DATA_BLOCK "MessagePrefix"   // DB31604
TITLE = CPG_MessagePrefix
{ S7_Optimized_Access := 'TRUE' }
AUTHOR : tech.team.motioncontrol@siemens.com
FAMILY : CPG
VERSION : 1.0
// Support: tech.team.motioncontrol@siemens.com
// Fax: +49 (0) 9131/98-1297
   VAR
      UN : Struct   // MessagePrefix for Unit
         Alarm : "CPG_typeMessagePrefix";   // MessagePrefix for Unit Alarms
      END_STRUCT;
      EM00 : Struct   // MessagePrefix for EquipmentModuleEM00
         EventControl : "CPG_typeMessagePrefix";   // MessagePrefixforEventControl
         CM01 : "CPG_typeMessagePrefix";   // MessagePrefixforControlModule#01
         CM02 : "CPG_typeMessagePrefix";   // MessagePrefixforControlModule#02
         CM03 : "CPG_typeMessagePrefix";   // MessagePrefixforControlModule#03
         CM04 : "CPG_typeMessagePrefix";   // MessagePrefixforControlModule#04
         CM05 : "CPG_typeMessagePrefix";   // MessagePrefixforControlModule#05
         CM06 : "CPG_typeMessagePrefix";   // MessagePrefixforControlModule#06
         CM07 : "CPG_typeMessagePrefix";   // MessagePrefixforControlModule#07
         CM08 : "CPG_typeMessagePrefix";   // MessagePrefixforControlModule#08
         CM09 : "CPG_typeMessagePrefix";   // MessagePrefixforControlModule#09
         CM10 : "CPG_typeMessagePrefix";   // MessagePrefixforControlModule#10
      END_STRUCT;
      EM01 : Struct   // MessagePrefix for EquipmentModuleEM01
         EventControl : "CPG_typeMessagePrefix";   // MessagePrefixforEventControl
         CM01 : "CPG_typeMessagePrefix";   // MessagePrefixforControlModule#01
         CM02 : "CPG_typeMessagePrefix";   // MessagePrefixforControlModule#02
         CM03 : "CPG_typeMessagePrefix";   // MessagePrefixforControlModule#03
         CM04 : "CPG_typeMessagePrefix";   // MessagePrefixforControlModule#04
         CM05 : "CPG_typeMessagePrefix";   // MessagePrefixforControlModule#05
         CM06 : "CPG_typeMessagePrefix";   // MessagePrefixforControlModule#06
         CM07 : "CPG_typeMessagePrefix";   // MessagePrefixforControlModule#07
         CM08 : "CPG_typeMessagePrefix";   // MessagePrefixforControlModule#08
         CM09 : "CPG_typeMessagePrefix";   // MessagePrefixforControlModule#09
         CM10 : "CPG_typeMessagePrefix";   // MessagePrefixforControlModule#10
      END_STRUCT;
      EM02 : Struct   // MessagePrefix for EquipmentModuleEM02
         EventControl : "CPG_typeMessagePrefix";   // MessagePrefixforEventControl
         CM01 : "CPG_typeMessagePrefix";   // MessagePrefixforControlModule#01
         CM02 : "CPG_typeMessagePrefix";   // MessagePrefixforControlModule#02
         CM03 : "CPG_typeMessagePrefix";   // MessagePrefixforControlModule#03
         CM04 : "CPG_typeMessagePrefix";   // MessagePrefixforControlModule#04
         CM05 : "CPG_typeMessagePrefix";   // MessagePrefixforControlModule#05
         CM06 : "CPG_typeMessagePrefix";   // MessagePrefixforControlModule#06
         CM07 : "CPG_typeMessagePrefix";   // MessagePrefixforControlModule#07
         CM08 : "CPG_typeMessagePrefix";   // MessagePrefixforControlModule#08
         CM09 : "CPG_typeMessagePrefix";   // MessagePrefixforControlModule#09
         CM10 : "CPG_typeMessagePrefix";   // MessagePrefixforControlModule#10
      END_STRUCT;
      EM03 : Struct   // MessagePrefix for EquipmentModuleEM03
         EventControl : "CPG_typeMessagePrefix";   // MessagePrefixforEventControl
         CM01 : "CPG_typeMessagePrefix";   // MessagePrefixforControlModule#01
         CM02 : "CPG_typeMessagePrefix";   // MessagePrefixforControlModule#02
         CM03 : "CPG_typeMessagePrefix";   // MessagePrefixforControlModule#03
         CM04 : "CPG_typeMessagePrefix";   // MessagePrefixforControlModule#04
         CM05 : "CPG_typeMessagePrefix";   // MessagePrefixforControlModule#05
         CM06 : "CPG_typeMessagePrefix";   // MessagePrefixforControlModule#06
         CM07 : "CPG_typeMessagePrefix";   // MessagePrefixforControlModule#07
         CM08 : "CPG_typeMessagePrefix";   // MessagePrefixforControlModule#08
         CM09 : "CPG_typeMessagePrefix";   // MessagePrefixforControlModule#09
         CM10 : "CPG_typeMessagePrefix";   // MessagePrefixforControlModule#10
      END_STRUCT;
      EM04 : Struct   // MessagePrefix for EquipmentModuleEM04
         EventControl : "CPG_typeMessagePrefix";   // MessagePrefixforEventControl
         CM01 : "CPG_typeMessagePrefix";   // MessagePrefixforControlModule#01
         CM02 : "CPG_typeMessagePrefix";   // MessagePrefixforControlModule#02
         CM03 : "CPG_typeMessagePrefix";   // MessagePrefixforControlModule#03
         CM04 : "CPG_typeMessagePrefix";   // MessagePrefixforControlModule#04
         CM05 : "CPG_typeMessagePrefix";   // MessagePrefixforControlModule#05
         CM06 : "CPG_typeMessagePrefix";   // MessagePrefixforControlModule#06
         CM07 : "CPG_typeMessagePrefix";   // MessagePrefixforControlModule#07
         CM08 : "CPG_typeMessagePrefix";   // MessagePrefixforControlModule#08
         CM09 : "CPG_typeMessagePrefix";   // MessagePrefixforControlModule#09
         CM10 : "CPG_typeMessagePrefix";   // MessagePrefixforControlModule#10
      END_STRUCT;
      EM05 : Struct   // MessagePrefix for EquipmentModuleEM05
         EventControl : "CPG_typeMessagePrefix";   // MessagePrefixforEventControl
         CM01 : "CPG_typeMessagePrefix";   // MessagePrefixforControlModule#01
         CM02 : "CPG_typeMessagePrefix";   // MessagePrefixforControlModule#02
         CM03 : "CPG_typeMessagePrefix";   // MessagePrefixforControlModule#03
         CM04 : "CPG_typeMessagePrefix";   // MessagePrefixforControlModule#04
         CM05 : "CPG_typeMessagePrefix";   // MessagePrefixforControlModule#05
         CM06 : "CPG_typeMessagePrefix";   // MessagePrefixforControlModule#06
         CM07 : "CPG_typeMessagePrefix";   // MessagePrefixforControlModule#07
         CM08 : "CPG_typeMessagePrefix";   // MessagePrefixforControlModule#08
         CM09 : "CPG_typeMessagePrefix";   // MessagePrefixforControlModule#09
         CM10 : "CPG_typeMessagePrefix";   // MessagePrefixforControlModule#10
      END_STRUCT;
      EM06 : Struct   // MessagePrefix for EquipmentModuleEM06
         EventControl : "CPG_typeMessagePrefix";   // MessagePrefixforEventControl
         CM01 : "CPG_typeMessagePrefix";   // MessagePrefixforControlModule#01
         CM02 : "CPG_typeMessagePrefix";   // MessagePrefixforControlModule#02
         CM03 : "CPG_typeMessagePrefix";   // MessagePrefixforControlModule#03
         CM04 : "CPG_typeMessagePrefix";   // MessagePrefixforControlModule#04
         CM05 : "CPG_typeMessagePrefix";   // MessagePrefixforControlModule#05
         CM06 : "CPG_typeMessagePrefix";   // MessagePrefixforControlModule#06
         CM07 : "CPG_typeMessagePrefix";   // MessagePrefixforControlModule#07
         CM08 : "CPG_typeMessagePrefix";   // MessagePrefixforControlModule#08
         CM09 : "CPG_typeMessagePrefix";   // MessagePrefixforControlModule#09
         CM10 : "CPG_typeMessagePrefix";   // MessagePrefixforControlModule#10
      END_STRUCT;
      EM07 : Struct   // MessagePrefix for EquipmentModuleEM07
         EventControl : "CPG_typeMessagePrefix";   // MessagePrefixforEventControl
         CM01 : "CPG_typeMessagePrefix";   // MessagePrefixforControlModule#01
         CM02 : "CPG_typeMessagePrefix";   // MessagePrefixforControlModule#02
         CM03 : "CPG_typeMessagePrefix";   // MessagePrefixforControlModule#03
         CM04 : "CPG_typeMessagePrefix";   // MessagePrefixforControlModule#04
         CM05 : "CPG_typeMessagePrefix";   // MessagePrefixforControlModule#05
         CM06 : "CPG_typeMessagePrefix";   // MessagePrefixforControlModule#06
         CM07 : "CPG_typeMessagePrefix";   // MessagePrefixforControlModule#07
         CM08 : "CPG_typeMessagePrefix";   // MessagePrefixforControlModule#08
         CM09 : "CPG_typeMessagePrefix";   // MessagePrefixforControlModule#09
         CM10 : "CPG_typeMessagePrefix";   // MessagePrefixforControlModule#10
      END_STRUCT;
      EM08 : Struct   // MessagePrefix for EquipmentModuleEM08
         EventControl : "CPG_typeMessagePrefix";   // MessagePrefixforEventControl
         CM01 : "CPG_typeMessagePrefix";   // MessagePrefixforControlModule#01
         CM02 : "CPG_typeMessagePrefix";   // MessagePrefixforControlModule#02
         CM03 : "CPG_typeMessagePrefix";   // MessagePrefixforControlModule#03
         CM04 : "CPG_typeMessagePrefix";   // MessagePrefixforControlModule#04
         CM05 : "CPG_typeMessagePrefix";   // MessagePrefixforControlModule#05
         CM06 : "CPG_typeMessagePrefix";   // MessagePrefixforControlModule#06
         CM07 : "CPG_typeMessagePrefix";   // MessagePrefixforControlModule#07
         CM08 : "CPG_typeMessagePrefix";   // MessagePrefixforControlModule#08
         CM09 : "CPG_typeMessagePrefix";   // MessagePrefixforControlModule#09
         CM10 : "CPG_typeMessagePrefix";   // MessagePrefixforControlModule#10
      END_STRUCT;
      EM09 : Struct   // MessagePrefix for EquipmentModuleEM09
         EventControl : "CPG_typeMessagePrefix";   // MessagePrefixforEventControl
         CM01 : "CPG_typeMessagePrefix";   // MessagePrefixforControlModule#01
         CM02 : "CPG_typeMessagePrefix";   // MessagePrefixforControlModule#02
         CM03 : "CPG_typeMessagePrefix";   // MessagePrefixforControlModule#03
         CM04 : "CPG_typeMessagePrefix";   // MessagePrefixforControlModule#04
         CM05 : "CPG_typeMessagePrefix";   // MessagePrefixforControlModule#05
         CM06 : "CPG_typeMessagePrefix";   // MessagePrefixforControlModule#06
         CM07 : "CPG_typeMessagePrefix";   // MessagePrefixforControlModule#07
         CM08 : "CPG_typeMessagePrefix";   // MessagePrefixforControlModule#08
         CM09 : "CPG_typeMessagePrefix";   // MessagePrefixforControlModule#09
         CM10 : "CPG_typeMessagePrefix";   // MessagePrefixforControlModule#10
      END_STRUCT;
   END_VAR
BEGIN
   UN.Alarm.messagePrefix[0] := 'Unit ';
   UN.Alarm.messagePrefix[1] := 'Unit ';
   EM00.EventControl.messagePrefix[0] := 'EM00 ';
   EM00.EventControl.messagePrefix[1] := 'EM00 ';
   EM00.CM01.messagePrefix[0] := 'CM01 ';
   EM00.CM01.messagePrefix[1] := 'CM01 ';
   EM00.CM02.messagePrefix[0] := 'CM02 ';
   EM00.CM02.messagePrefix[1] := 'CM02 ';
   EM00.CM03.messagePrefix[0] := 'CM03 ';
   EM00.CM03.messagePrefix[1] := 'CM03 ';
   EM00.CM04.messagePrefix[0] := 'CM04 ';
   EM00.CM04.messagePrefix[1] := 'CM04 ';
   EM00.CM05.messagePrefix[0] := 'CM05 ';
   EM00.CM05.messagePrefix[1] := 'CM05 ';
   EM00.CM06.messagePrefix[0] := 'CM06 ';
   EM00.CM06.messagePrefix[1] := 'CM06 ';
   EM00.CM07.messagePrefix[0] := 'CM07 ';
   EM00.CM07.messagePrefix[1] := 'CM07 ';
   EM00.CM08.messagePrefix[0] := 'CM08 ';
   EM00.CM08.messagePrefix[1] := 'CM08 ';
   EM00.CM09.messagePrefix[0] := 'CM09 ';
   EM00.CM09.messagePrefix[1] := 'CM09 ';
   EM00.CM10.messagePrefix[0] := 'CM10 ';
   EM00.CM10.messagePrefix[1] := 'CM10 ';
   EM09.CM10.messagePrefix[1] := 'CM10 ';
   EM09.CM10.messagePrefix[0] := 'CM10 ';
   EM09.CM09.messagePrefix[1] := 'CM09 ';
   EM09.CM09.messagePrefix[0] := 'CM09 ';
   EM09.CM08.messagePrefix[1] := 'CM08 ';
   EM09.CM08.messagePrefix[0] := 'CM08 ';
   EM09.CM07.messagePrefix[1] := 'CM07 ';
   EM09.CM07.messagePrefix[0] := 'CM07 ';
   EM09.CM06.messagePrefix[1] := 'CM06 ';
   EM09.CM06.messagePrefix[0] := 'CM06 ';
   EM09.CM05.messagePrefix[1] := 'CM05 ';
   EM09.CM05.messagePrefix[0] := 'CM05 ';
   EM09.CM04.messagePrefix[1] := 'CM04 ';
   EM09.CM04.messagePrefix[0] := 'CM04 ';
   EM09.CM03.messagePrefix[1] := 'CM03 ';
   EM09.CM03.messagePrefix[0] := 'CM03 ';
   EM09.CM02.messagePrefix[1] := 'CM02 ';
   EM09.CM02.messagePrefix[0] := 'CM02 ';
   EM09.CM01.messagePrefix[1] := 'CM01 ';
   EM09.CM01.messagePrefix[0] := 'CM01 ';
   EM09.EventControl.messagePrefix[1] := 'EM09 ';
   EM09.EventControl.messagePrefix[0] := 'EM09 ';
   EM08.CM10.messagePrefix[1] := 'CM10 ';
   EM08.CM10.messagePrefix[0] := 'CM10 ';
   EM08.CM09.messagePrefix[1] := 'CM09 ';
   EM08.CM09.messagePrefix[0] := 'CM09 ';
   EM08.CM08.messagePrefix[1] := 'CM08 ';
   EM08.CM08.messagePrefix[0] := 'CM08 ';
   EM08.CM07.messagePrefix[1] := 'CM07 ';
   EM08.CM07.messagePrefix[0] := 'CM07 ';
   EM08.CM06.messagePrefix[1] := 'CM06 ';
   EM08.CM06.messagePrefix[0] := 'CM06 ';
   EM08.CM05.messagePrefix[1] := 'CM05 ';
   EM08.CM05.messagePrefix[0] := 'CM05 ';
   EM08.CM04.messagePrefix[1] := 'CM04 ';
   EM08.CM04.messagePrefix[0] := 'CM04 ';
   EM08.CM03.messagePrefix[1] := 'CM03 ';
   EM08.CM03.messagePrefix[0] := 'CM03 ';
   EM08.CM02.messagePrefix[1] := 'CM02 ';
   EM08.CM02.messagePrefix[0] := 'CM02 ';
   EM08.CM01.messagePrefix[1] := 'CM01 ';
   EM08.CM01.messagePrefix[0] := 'CM01 ';
   EM08.EventControl.messagePrefix[1] := 'EM08 ';
   EM08.EventControl.messagePrefix[0] := 'EM08 ';
   EM07.CM10.messagePrefix[1] := 'CM10 ';
   EM07.CM10.messagePrefix[0] := 'CM10 ';
   EM07.CM09.messagePrefix[1] := 'CM09 ';
   EM07.CM09.messagePrefix[0] := 'CM09 ';
   EM07.CM08.messagePrefix[1] := 'CM08 ';
   EM07.CM08.messagePrefix[0] := 'CM08 ';
   EM07.CM07.messagePrefix[1] := 'CM07 ';
   EM07.CM07.messagePrefix[0] := 'CM07 ';
   EM07.CM06.messagePrefix[1] := 'CM06 ';
   EM07.CM06.messagePrefix[0] := 'CM06 ';
   EM07.CM05.messagePrefix[1] := 'CM05 ';
   EM07.CM05.messagePrefix[0] := 'CM05 ';
   EM07.CM04.messagePrefix[1] := 'CM04 ';
   EM07.CM04.messagePrefix[0] := 'CM04 ';
   EM07.CM03.messagePrefix[1] := 'CM03 ';
   EM07.CM03.messagePrefix[0] := 'CM03 ';
   EM07.CM02.messagePrefix[1] := 'CM02 ';
   EM07.CM02.messagePrefix[0] := 'CM02 ';
   EM07.CM01.messagePrefix[1] := 'CM01 ';
   EM07.CM01.messagePrefix[0] := 'CM01 ';
   EM07.EventControl.messagePrefix[1] := 'EM07 ';
   EM07.EventControl.messagePrefix[0] := 'EM07 ';
   EM06.CM10.messagePrefix[1] := 'CM10 ';
   EM06.CM10.messagePrefix[0] := 'CM10 ';
   EM06.CM09.messagePrefix[1] := 'CM09 ';
   EM06.CM09.messagePrefix[0] := 'CM09 ';
   EM06.CM08.messagePrefix[1] := 'CM08 ';
   EM06.CM08.messagePrefix[0] := 'CM08 ';
   EM06.CM07.messagePrefix[1] := 'CM07 ';
   EM06.CM07.messagePrefix[0] := 'CM07 ';
   EM06.CM06.messagePrefix[1] := 'CM06 ';
   EM06.CM06.messagePrefix[0] := 'CM06 ';
   EM06.CM05.messagePrefix[1] := 'CM05 ';
   EM06.CM05.messagePrefix[0] := 'CM05 ';
   EM06.CM04.messagePrefix[1] := 'CM04 ';
   EM06.CM04.messagePrefix[0] := 'CM04 ';
   EM06.CM03.messagePrefix[1] := 'CM03 ';
   EM06.CM03.messagePrefix[0] := 'CM03 ';
   EM06.CM02.messagePrefix[1] := 'CM02 ';
   EM06.CM02.messagePrefix[0] := 'CM02 ';
   EM06.CM01.messagePrefix[1] := 'CM01 ';
   EM06.CM01.messagePrefix[0] := 'CM01 ';
   EM06.EventControl.messagePrefix[1] := 'EM06 ';
   EM06.EventControl.messagePrefix[0] := 'EM06 ';
   EM05.CM10.messagePrefix[1] := 'CM10 ';
   EM05.CM10.messagePrefix[0] := 'CM10 ';
   EM05.CM09.messagePrefix[1] := 'CM09 ';
   EM05.CM09.messagePrefix[0] := 'CM09 ';
   EM05.CM08.messagePrefix[1] := 'CM08 ';
   EM05.CM08.messagePrefix[0] := 'CM08 ';
   EM05.CM07.messagePrefix[1] := 'CM07 ';
   EM05.CM07.messagePrefix[0] := 'CM07 ';
   EM05.CM06.messagePrefix[1] := 'CM06 ';
   EM05.CM06.messagePrefix[0] := 'CM06 ';
   EM05.CM05.messagePrefix[1] := 'CM05 ';
   EM05.CM05.messagePrefix[0] := 'CM05 ';
   EM05.CM04.messagePrefix[1] := 'CM04 ';
   EM05.CM04.messagePrefix[0] := 'CM04 ';
   EM05.CM03.messagePrefix[1] := 'CM03 ';
   EM05.CM03.messagePrefix[0] := 'CM03 ';
   EM05.CM02.messagePrefix[1] := 'CM02 ';
   EM05.CM02.messagePrefix[0] := 'CM02 ';
   EM05.CM01.messagePrefix[1] := 'CM01 ';
   EM05.CM01.messagePrefix[0] := 'CM01 ';
   EM05.EventControl.messagePrefix[1] := 'EM05 ';
   EM05.EventControl.messagePrefix[0] := 'EM05 ';
   EM04.CM10.messagePrefix[1] := 'CM10 ';
   EM04.CM10.messagePrefix[0] := 'CM10 ';
   EM04.CM09.messagePrefix[1] := 'CM09 ';
   EM04.CM09.messagePrefix[0] := 'CM09 ';
   EM04.CM08.messagePrefix[1] := 'CM08 ';
   EM04.CM08.messagePrefix[0] := 'CM08 ';
   EM04.CM07.messagePrefix[1] := 'CM07 ';
   EM04.CM07.messagePrefix[0] := 'CM07 ';
   EM04.CM06.messagePrefix[1] := 'CM06 ';
   EM04.CM06.messagePrefix[0] := 'CM06 ';
   EM04.CM05.messagePrefix[1] := 'CM05 ';
   EM04.CM05.messagePrefix[0] := 'CM05 ';
   EM04.CM04.messagePrefix[1] := 'CM04 ';
   EM04.CM04.messagePrefix[0] := 'CM04 ';
   EM04.CM03.messagePrefix[1] := 'CM03 ';
   EM04.CM03.messagePrefix[0] := 'CM03 ';
   EM04.CM02.messagePrefix[1] := 'CM02 ';
   EM04.CM02.messagePrefix[0] := 'CM02 ';
   EM04.CM01.messagePrefix[1] := 'CM01 ';
   EM04.CM01.messagePrefix[0] := 'CM01 ';
   EM04.EventControl.messagePrefix[1] := 'EM04 ';
   EM04.EventControl.messagePrefix[0] := 'EM04 ';
   EM03.CM10.messagePrefix[1] := 'CM10 ';
   EM03.CM10.messagePrefix[0] := 'CM10 ';
   EM03.CM09.messagePrefix[1] := 'CM09 ';
   EM03.CM09.messagePrefix[0] := 'CM09 ';
   EM03.CM08.messagePrefix[1] := 'CM08 ';
   EM03.CM08.messagePrefix[0] := 'CM08 ';
   EM03.CM07.messagePrefix[1] := 'CM07 ';
   EM03.CM07.messagePrefix[0] := 'CM07 ';
   EM03.CM06.messagePrefix[1] := 'CM06 ';
   EM03.CM06.messagePrefix[0] := 'CM06 ';
   EM03.CM05.messagePrefix[1] := 'CM05 ';
   EM03.CM05.messagePrefix[0] := 'CM05 ';
   EM03.CM04.messagePrefix[1] := 'CM04 ';
   EM03.CM04.messagePrefix[0] := 'CM04 ';
   EM03.CM03.messagePrefix[1] := 'CM03 ';
   EM03.CM03.messagePrefix[0] := 'CM03 ';
   EM03.CM02.messagePrefix[1] := 'CM02 ';
   EM03.CM02.messagePrefix[0] := 'CM02 ';
   EM03.CM01.messagePrefix[1] := 'CM01 ';
   EM03.CM01.messagePrefix[0] := 'CM01 ';
   EM03.EventControl.messagePrefix[1] := 'EM03 ';
   EM03.EventControl.messagePrefix[0] := 'EM03 ';
   EM02.CM10.messagePrefix[1] := 'CM10 ';
   EM02.CM10.messagePrefix[0] := 'CM10 ';
   EM02.CM09.messagePrefix[1] := 'CM09 ';
   EM02.CM09.messagePrefix[0] := 'CM09 ';
   EM02.CM08.messagePrefix[1] := 'CM08 ';
   EM02.CM08.messagePrefix[0] := 'CM08 ';
   EM02.CM07.messagePrefix[1] := 'CM07 ';
   EM02.CM07.messagePrefix[0] := 'CM07 ';
   EM02.CM06.messagePrefix[1] := 'CM06 ';
   EM02.CM06.messagePrefix[0] := 'CM06 ';
   EM02.CM05.messagePrefix[1] := 'CM05 ';
   EM02.CM05.messagePrefix[0] := 'CM05 ';
   EM02.CM04.messagePrefix[1] := 'CM04 ';
   EM02.CM04.messagePrefix[0] := 'CM04 ';
   EM02.CM03.messagePrefix[1] := 'CM03 ';
   EM02.CM03.messagePrefix[0] := 'CM03 ';
   EM02.CM02.messagePrefix[1] := 'CM02 ';
   EM02.CM02.messagePrefix[0] := 'CM02 ';
   EM02.CM01.messagePrefix[1] := 'CM01 ';
   EM02.CM01.messagePrefix[0] := 'CM01 ';
   EM02.EventControl.messagePrefix[1] := 'EM01 ';
   EM02.EventControl.messagePrefix[0] := 'EM01 ';
   EM01.CM10.messagePrefix[1] := 'CM10 ';
   EM01.CM10.messagePrefix[0] := 'CM10 ';
   EM01.CM09.messagePrefix[1] := 'CM09 ';
   EM01.CM09.messagePrefix[0] := 'CM09 ';
   EM01.CM08.messagePrefix[1] := 'CM08 ';
   EM01.CM08.messagePrefix[0] := 'CM08 ';
   EM01.CM07.messagePrefix[1] := 'CM07 ';
   EM01.CM07.messagePrefix[0] := 'CM07 ';
   EM01.CM06.messagePrefix[1] := 'CM06 ';
   EM01.CM06.messagePrefix[0] := 'CM06 ';
   EM01.CM05.messagePrefix[1] := 'CM05 ';
   EM01.CM05.messagePrefix[0] := 'CM05 ';
   EM01.CM04.messagePrefix[1] := 'CM04 ';
   EM01.CM04.messagePrefix[0] := 'CM04 ';
   EM01.CM03.messagePrefix[1] := 'CM03 ';
   EM01.CM03.messagePrefix[0] := 'CM03 ';
   EM01.CM02.messagePrefix[1] := 'CM02 ';
   EM01.CM02.messagePrefix[0] := 'CM02 ';
   EM01.CM01.messagePrefix[1] := 'CM01 ';
   EM01.CM01.messagePrefix[0] := 'CM01 ';
   EM01.EventControl.messagePrefix[1] := 'EM01 ';
   EM01.EventControl.messagePrefix[0] := 'EM01 ';
   UN.Alarm.messagePrefix[2] := 'Unit ';
   EM00.EventControl.messagePrefix[2] := 'EM00 ';
   EM00.CM01.messagePrefix[2] := 'CM01 ';
   EM00.CM02.messagePrefix[2] := 'CM02 ';
   EM00.CM03.messagePrefix[2] := 'CM03 ';
   EM00.CM04.messagePrefix[2] := 'CM04 ';
   EM00.CM05.messagePrefix[2] := 'CM05 ';
   EM00.CM06.messagePrefix[2] := 'CM06 ';
   EM00.CM07.messagePrefix[2] := 'CM07 ';
   EM00.CM08.messagePrefix[2] := 'CM08 ';
   EM00.CM09.messagePrefix[2] := 'CM09 ';
   EM00.CM10.messagePrefix[2] := 'CM10 ';
   EM01.EventControl.messagePrefix[2] := 'EM01 ';
   EM01.CM01.messagePrefix[2] := 'CM01 ';
   EM01.CM02.messagePrefix[2] := 'CM02 ';
   EM01.CM03.messagePrefix[2] := 'CM03 ';
   EM01.CM04.messagePrefix[2] := 'CM04 ';
   EM01.CM05.messagePrefix[2] := 'CM05 ';
   EM01.CM06.messagePrefix[2] := 'CM06 ';
   EM01.CM07.messagePrefix[2] := 'CM07 ';
   EM01.CM08.messagePrefix[2] := 'CM08 ';
   EM01.CM09.messagePrefix[2] := 'CM09 ';
   EM01.CM10.messagePrefix[2] := 'CM10 ';
   EM02.EventControl.messagePrefix[2] := 'EM01 ';
   EM02.CM01.messagePrefix[2] := 'CM01 ';
   EM02.CM02.messagePrefix[2] := 'CM02 ';
   EM02.CM03.messagePrefix[2] := 'CM03 ';
   EM02.CM04.messagePrefix[2] := 'CM04 ';
   EM02.CM05.messagePrefix[2] := 'CM05 ';
   EM02.CM06.messagePrefix[2] := 'CM06 ';
   EM02.CM07.messagePrefix[2] := 'CM07 ';
   EM02.CM08.messagePrefix[2] := 'CM08 ';
   EM02.CM09.messagePrefix[2] := 'CM09 ';
   EM02.CM10.messagePrefix[2] := 'CM10 ';
   EM03.EventControl.messagePrefix[2] := 'EM03 ';
   EM03.CM01.messagePrefix[2] := 'CM01 ';
   EM03.CM02.messagePrefix[2] := 'CM02 ';
   EM03.CM03.messagePrefix[2] := 'CM03 ';
   EM03.CM04.messagePrefix[2] := 'CM04 ';
   EM03.CM05.messagePrefix[2] := 'CM05 ';
   EM03.CM06.messagePrefix[2] := 'CM06 ';
   EM03.CM07.messagePrefix[2] := 'CM07 ';
   EM03.CM08.messagePrefix[2] := 'CM08 ';
   EM03.CM09.messagePrefix[2] := 'CM09 ';
   EM03.CM10.messagePrefix[2] := 'CM10 ';
   EM04.EventControl.messagePrefix[2] := 'EM04 ';
   EM04.CM01.messagePrefix[2] := 'CM01 ';
   EM04.CM02.messagePrefix[2] := 'CM02 ';
   EM04.CM03.messagePrefix[2] := 'CM03 ';
   EM04.CM04.messagePrefix[2] := 'CM04 ';
   EM04.CM05.messagePrefix[2] := 'CM05 ';
   EM04.CM06.messagePrefix[2] := 'CM06 ';
   EM04.CM07.messagePrefix[2] := 'CM07 ';
   EM04.CM08.messagePrefix[2] := 'CM08 ';
   EM04.CM09.messagePrefix[2] := 'CM09 ';
   EM04.CM10.messagePrefix[2] := 'CM10 ';
   EM05.EventControl.messagePrefix[2] := 'EM05 ';
   EM05.CM01.messagePrefix[2] := 'CM01 ';
   EM05.CM02.messagePrefix[2] := 'CM02 ';
   EM05.CM03.messagePrefix[2] := 'CM03 ';
   EM05.CM04.messagePrefix[2] := 'CM04 ';
   EM05.CM05.messagePrefix[2] := 'CM05 ';
   EM05.CM06.messagePrefix[2] := 'CM06 ';
   EM05.CM07.messagePrefix[2] := 'CM07 ';
   EM05.CM08.messagePrefix[2] := 'CM08 ';
   EM05.CM09.messagePrefix[2] := 'CM09 ';
   EM05.CM10.messagePrefix[2] := 'CM10 ';
   EM06.EventControl.messagePrefix[2] := 'EM06 ';
   EM06.CM01.messagePrefix[2] := 'CM01 ';
   EM06.CM02.messagePrefix[2] := 'CM02 ';
   EM06.CM03.messagePrefix[2] := 'CM03 ';
   EM06.CM04.messagePrefix[2] := 'CM04 ';
   EM06.CM05.messagePrefix[2] := 'CM05 ';
   EM06.CM06.messagePrefix[2] := 'CM06 ';
   EM06.CM07.messagePrefix[2] := 'CM07 ';
   EM06.CM08.messagePrefix[2] := 'CM08 ';
   EM06.CM09.messagePrefix[2] := 'CM09 ';
   EM06.CM10.messagePrefix[2] := 'CM10 ';
   EM07.EventControl.messagePrefix[2] := 'EM07 ';
   EM07.CM01.messagePrefix[2] := 'CM01 ';
   EM07.CM02.messagePrefix[2] := 'CM02 ';
   EM07.CM03.messagePrefix[2] := 'CM03 ';
   EM07.CM04.messagePrefix[2] := 'CM04 ';
   EM07.CM05.messagePrefix[2] := 'CM05 ';
   EM07.CM06.messagePrefix[2] := 'CM06 ';
   EM07.CM07.messagePrefix[2] := 'CM07 ';
   EM07.CM08.messagePrefix[2] := 'CM08 ';
   EM07.CM09.messagePrefix[2] := 'CM09 ';
   EM07.CM10.messagePrefix[2] := 'CM10 ';
   EM08.EventControl.messagePrefix[2] := 'EM08 ';
   EM08.CM01.messagePrefix[2] := 'CM01 ';
   EM08.CM02.messagePrefix[2] := 'CM02 ';
   EM08.CM03.messagePrefix[2] := 'CM03 ';
   EM08.CM04.messagePrefix[2] := 'CM04 ';
   EM08.CM05.messagePrefix[2] := 'CM05 ';
   EM08.CM06.messagePrefix[2] := 'CM06 ';
   EM08.CM07.messagePrefix[2] := 'CM07 ';
   EM08.CM08.messagePrefix[2] := 'CM08 ';
   EM08.CM09.messagePrefix[2] := 'CM09 ';
   EM08.CM10.messagePrefix[2] := 'CM10 ';
   EM09.EventControl.messagePrefix[2] := 'EM09 ';
   EM09.CM01.messagePrefix[2] := 'CM01 ';
   EM09.CM02.messagePrefix[2] := 'CM02 ';
   EM09.CM03.messagePrefix[2] := 'CM03 ';
   EM09.CM04.messagePrefix[2] := 'CM04 ';
   EM09.CM05.messagePrefix[2] := 'CM05 ';
   EM09.CM06.messagePrefix[2] := 'CM06 ';
   EM09.CM07.messagePrefix[2] := 'CM07 ';
   EM09.CM08.messagePrefix[2] := 'CM08 ';
   EM09.CM09.messagePrefix[2] := 'CM09 ';
   EM09.CM10.messagePrefix[2] := 'CM10 ';
END_DATA_BLOCK

// folder: SupportingBlocks/CPG_Blocks

DATA_BLOCK "WarningCfg"   // DB31601
TITLE = CPG_WarningCfg
{ S7_Optimized_Access := 'TRUE' }
AUTHOR : tech.team.motioncontrol@siemens.com
FAMILY : CPG
VERSION : 1.0
// Support: tech.team.motioncontrol@siemens.com
// Fax: +49 (0) 9131/98-1297
   VAR
      Event : Array[0.."CPG_NO_OF_CFG_WARNINGS_UPPER_LIM"] of "CPG_typeEventCfg";
   END_VAR
BEGIN
   Event[0].message[0] := 'Warning Test';
   Event[0].message[1] := 'Warning Test';
   Event[1].message[0] := 'Low Bottle Supply';
   Event[1].message[1] := 'Flaschenzufuhr niedrig';
   Event[2].message[0] := 'Low Label Supply';
   Event[2].message[1] := 'Etikettenzufuhr niedrig';
   Event[29].message[1] := 'Reserve';
   Event[29].message[0] := 'Spare';
   Event[28].message[1] := 'Reserve';
   Event[28].message[0] := 'Spare';
   Event[27].message[1] := 'Reserve';
   Event[27].message[0] := 'Spare';
   Event[26].message[1] := 'Reserve';
   Event[26].message[0] := 'Spare';
   Event[25].message[0] := 'Spare';
   Event[25].message[1] := 'Reserve';
   Event[24].message[0] := 'Spare';
   Event[24].message[1] := 'Reserve';
   Event[23].message[0] := 'Spare';
   Event[23].message[1] := 'Reserve';
   Event[22].message[0] := 'Spare';
   Event[22].message[1] := 'Reserve';
   Event[21].message[0] := 'Spare';
   Event[21].message[1] := 'Reserve';
   Event[20].message[0] := 'Spare';
   Event[20].message[1] := 'Reserve';
   Event[19].message[0] := 'Spare';
   Event[19].message[1] := 'Reserve';
   Event[18].message[0] := 'Spare';
   Event[18].message[1] := 'Reserve';
   Event[17].message[0] := 'Spare';
   Event[17].message[1] := 'Reserve';
   Event[16].message[0] := 'Spare';
   Event[16].message[1] := 'Reserve';
   Event[15].message[0] := 'Spare';
   Event[15].message[1] := 'Reserve';
   Event[14].message[0] := 'Spare';
   Event[14].message[1] := 'Reserve';
   Event[13].message[0] := 'Spare';
   Event[13].message[1] := 'Reserve';
   Event[12].message[1] := 'Reserve';
   Event[12].message[0] := 'Spare';
   Event[11].message[1] := 'Reserve';
   Event[11].message[0] := 'Spare';
   Event[10].message[0] := 'Spare';
   Event[10].message[1] := 'Reserve';
   Event[9].message[0] := 'Spare';
   Event[9].message[1] := 'Reserve';
   Event[8].message[0] := 'Spare';
   Event[8].message[1] := 'Reserve';
   Event[7].message[0] := 'Spare';
   Event[7].message[1] := 'Reserve';
   Event[6].message[0] := 'Spare';
   Event[6].message[1] := 'Reserve';
   Event[5].message[0] := 'Spare';
   Event[5].message[1] := 'Reserve';
   Event[3].message[0] := 'Spare';
   Event[3].message[1] := 'Reserve';
   Event[4].message[1] := 'Reserve';
   Event[4].message[0] := 'Spare';
   Event[0].ID := 0;
   Event[1].ID := 1;
   Event[2].ID := 2;
   Event[3].ID := 3;
   Event[4].ID := 4;
   Event[5].ID := 5;
   Event[6].ID := 6;
   Event[7].ID := 7;
   Event[8].ID := 8;
   Event[9].ID := 9;
   Event[10].ID := 10;
   Event[11].ID := 11;
   Event[12].ID := 12;
   Event[13].ID := 13;
   Event[14].ID := 14;
   Event[15].ID := 15;
   Event[16].ID := 16;
   Event[17].ID := 17;
   Event[18].ID := 18;
   Event[19].ID := 19;
   Event[20].ID := 20;
   Event[21].ID := 21;
   Event[22].ID := 22;
   Event[23].ID := 23;
   Event[24].ID := 24;
   Event[25].ID := 25;
   Event[26].ID := 26;
   Event[27].ID := 27;
   Event[28].ID := 28;
   Event[29].ID := 29;
   Event[0].message[2] := 'Los Warning Test';
   Event[1].message[2] := 'Las Low Bottle Supply';
   Event[2].message[2] := 'Las Low Label Supply';
   Event[3].message[2] := 'Spare';
   Event[4].message[2] := 'Spare';
   Event[5].message[2] := 'Spare';
   Event[6].message[2] := 'Spare';
   Event[7].message[2] := 'Spare';
   Event[8].message[2] := 'Spare';
   Event[9].message[2] := 'Spare';
   Event[10].message[2] := 'Spare';
   Event[11].message[2] := 'Spare';
   Event[12].message[2] := 'Spare';
   Event[13].message[2] := 'Spare';
   Event[14].message[2] := 'Spare';
   Event[15].message[2] := 'Spare';
   Event[16].message[2] := 'Spare';
   Event[17].message[2] := 'Spare';
   Event[18].message[2] := 'Spare';
   Event[19].message[2] := 'Spare';
   Event[20].message[2] := 'Spare';
   Event[21].message[2] := 'Spare';
   Event[22].message[2] := 'Spare';
   Event[23].message[2] := 'Spare';
   Event[24].message[2] := 'Spare';
   Event[25].message[2] := 'Spare';
   Event[26].message[2] := 'Spare';
   Event[27].message[2] := 'Spare';
   Event[28].message[2] := 'Spare';
   Event[29].message[2] := 'Spare';
   // Event[0] : Warning Test
   // Event[1] : Low Bottle Supply
   // Event[2] : Low Label Supply
   // Event[3] : Spare
   // Event[4] : Spare
   // Event[5] : Spare
   // Event[6] : Spare
   // Event[7] : Spare
   // Event[8] : Spare
   // Event[9] : Spare
   // Event[10] : Spare
   // Event[11] : Spare
   // Event[12] : Spare
   // Event[13] : Spare
   // Event[14] : Spare
   // Event[15] : Spare
   // Event[16] : Spare
   // Event[17] : Spare
   // Event[18] : Spare
   // Event[19] : Spare
   // Event[20] : Spare
   // Event[21] : Spare
   // Event[22] : Spare
   // Event[23] : Spare
   // Event[24] : Spare
   // Event[25] : Spare
   // Event[26] : Spare
   // Event[27] : Spare
   // Event[28] : Spare
   // Event[29] : Spare
END_DATA_BLOCK

// folder: _UN01_Palletizer

DATA_BLOCK "UN"   // DB31629
TITLE = UN
{ S7_Optimized_Access := 'TRUE' }
AUTHOR : tech.team.motioncontrol@siemens.com
FAMILY : CPG
VERSION : 1.0
// Support: tech.team.motioncontrol@siemens.com
// Fax: +49 (0) 9131/98-1297
   VAR
      PackML_Sts : "CPG_typePackML_ModuleSts";   // PackML Module Status - UN Status
      PackML_Sts_Alarm : "CPG_typePackML_ModuleSts";   // PackML Module Status - UN alarm status
      Alarm : "CPG_typeEventStatus";   // Alarm Event Status - UN Status
      Warning : "CPG_typeEventStatus";   // Warning Event Status - UN Status
      Status : "CPG_typeEventStatus";   // Event Status - UN Status
   END_VAR
BEGIN
END_DATA_BLOCK

// folder: _UN01_Palletizer/Instances

DATA_BLOCK "InstUN_00_Main"   // DB31620
TITLE = instUN00_00_Main
{ S7_Optimized_Access := 'TRUE' }
AUTHOR : tech.team.motioncontrol@siemens.com
FAMILY : CPG
VERSION : 1.0
// Support: tech.team.motioncontrol@siemens.com
// Fax: +49 (0) 9131/98-1297
// stored: InstanceOfName UN_00_Main
"UN_00_Main"
BEGIN
END_DATA_BLOCK

// folder: (top level)

FUNCTION "MHJ-PLC-Lab-Function-S71500" : Void   // FC9000, SCL
{ S7_Optimized_Access := 'TRUE' }
VERSION : 0.1
   VAR_TEMP
      Value : Byte;
      ForCounter : Int;
   END_VAR
   VAR CONSTANT
      Value_01_DW : DWord := 16#1223_5486;
      Value_02_DW : DWord := 16#A6C9_D1F5;
   END_VAR
BEGIN

   #Value:=PEEK(area := 16#82,
        dbNumber := 0,
        byteOffset := 511);
   #Value := #Value + 1;

   POKE(area := 16#82,
        dbNumber := 0,
        byteOffset := 511,
        value := #Value);

   POKE(area := 16#82,
        dbNumber := 0,
        byteOffset := 1016,
        value := #Value_01_DW);
   POKE(area := 16#82,
        dbNumber := 0,
        byteOffset := 1020,
        value := #Value_02_DW);

   FOR #ForCounter := 0 TO 63 DO
       #Value:=PEEK(area := 16#1,
            dbNumber := 0,
            byteOffset := #ForCounter);
       POKE(area := 16#81,
            dbNumber := 0,
            byteOffset := #ForCounter,
            value := #Value);
   END_FOR;
   #Value := PEEK(area := 16#1,
                  dbNumber := 0,
                  byteOffset := 512);
   POKE(area := 16#82,
        dbNumber := 0,
        byteOffset := 512,
        value := #Value);
END_FUNCTION

ORGANIZATION_BLOCK "Main"   // OB1, LAD, ProgramCycle
TITLE = Main
{ S7_Optimized_Access := 'TRUE' }
AUTHOR : tech.team.motioncontrol@siemens.com
FAMILY : CPG
VERSION : 1.0
// Support: tech.team.motioncontrol@siemens.com
// Fax: +49 (0) 9131/98-1297
   VAR_INPUT
      Initial_Call : Bool;   // Initial call of this OB
      Remanence : Bool;   // =True, if remanent data are available
   END_VAR
   VAR_TEMP   // added for the SCL form of the ladder/FBD networks
      _w1 : Bool;
   END_VAR
BEGIN

REGION Network 1: Factory IO PLCSIM Communication
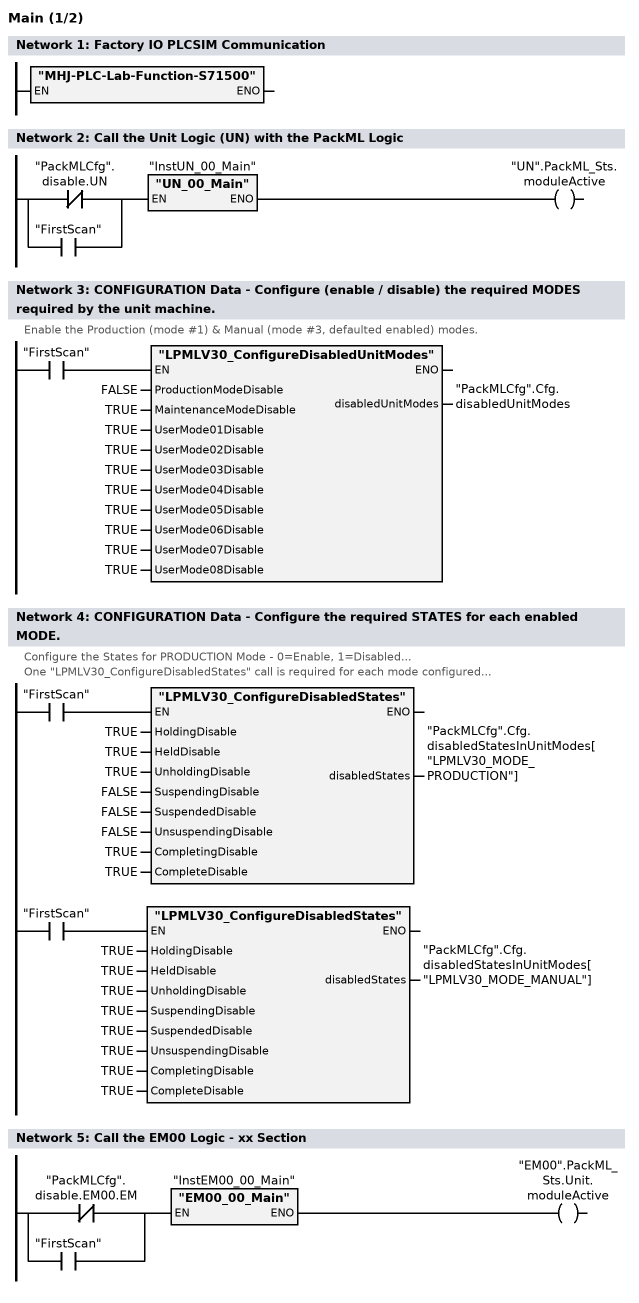
   RUNG wire#powerrail
      "MHJ-PLC-Lab-Function-S71500"()
   END_RUNG
   // the same network as SCL:
   "MHJ-PLC-Lab-Function-S71500"();
END_REGION

REGION Network 2: Call the Unit Logic (UN) with the PackML Logic
   RUNG wire#powerrail
      I_Contact( "PackMLCfg".disable.UN )
      wire#w1
      "InstUN_00_Main"()
      Coil( "UN".PackML_Sts.moduleActive )
   END_RUNG
   RUNG wire#powerrail
      Contact( "FirstScan" )
   END_RUNG wire#w1
   // the same network as SCL:
   "InstUN_00_Main"(EN := NOT "PackMLCfg".disable.UN OR "FirstScan", ENO => #_w1);   // "UN_00_Main"
   "UN".PackML_Sts.moduleActive := #_w1;
END_REGION

REGION Network 3: CONFIGURATION Data - Configure (enable / disable) the required MODES required by the unit machine.
   // Enable the Production (mode #1) & Manual (mode #3, defaulted enabled) modes.
   RUNG wire#powerrail
      Contact( "FirstScan" )
      "LPMLV30_ConfigureDisabledUnitModes"(ProductionModeDisable := FALSE, MaintenanceModeDisable := TRUE, UserMode01Disable := TRUE, UserMode02Disable := TRUE, UserMode03Disable := TRUE, UserMode04Disable := TRUE, UserMode05Disable := TRUE, UserMode06Disable := TRUE, UserMode07Disable := TRUE, UserMode08Disable := TRUE, disabledUnitModes => "PackMLCfg".Cfg.disabledUnitModes)
   END_RUNG
   // the same network as SCL:
   IF "FirstScan" THEN
       "LPMLV30_ConfigureDisabledUnitModes"(ProductionModeDisable := FALSE,
                               MaintenanceModeDisable := TRUE,
                               UserMode01Disable := TRUE,
                               UserMode02Disable := TRUE,
                               UserMode03Disable := TRUE,
                               UserMode04Disable := TRUE,
                               UserMode05Disable := TRUE,
                               UserMode06Disable := TRUE,
                               UserMode07Disable := TRUE,
                               UserMode08Disable := TRUE,
                               disabledUnitModes => "PackMLCfg".Cfg.disabledUnitModes);
   END_IF;
END_REGION

REGION Network 4: CONFIGURATION Data - Configure the required STATES for each enabled MODE.
   // Configure the States for PRODUCTION Mode - 0=Enable, 1=Disabled...
   // One "LPMLV30_ConfigureDisabledStates" call is required for each mode configured...
   RUNG wire#powerrail
      Contact( "FirstScan" )
      "LPMLV30_ConfigureDisabledStates"(HoldingDisable := TRUE, HeldDisable := TRUE, UnholdingDisable := TRUE, SuspendingDisable := FALSE, SuspendedDisable := FALSE, UnsuspendingDisable := FALSE, CompletingDisable := TRUE, CompleteDisable := TRUE, disabledStates => "PackMLCfg".Cfg.disabledStatesInUnitModes["LPMLV30_MODE_PRODUCTION"])
   END_RUNG
   RUNG wire#powerrail
      Contact( "FirstScan" )
      "LPMLV30_ConfigureDisabledStates"(HoldingDisable := TRUE, HeldDisable := TRUE, UnholdingDisable := TRUE, SuspendingDisable := TRUE, SuspendedDisable := TRUE, UnsuspendingDisable := TRUE, CompletingDisable := TRUE, CompleteDisable := TRUE, disabledStates => "PackMLCfg".Cfg.disabledStatesInUnitModes["LPMLV30_MODE_MANUAL"])
   END_RUNG
   // the same network as SCL:
   IF "FirstScan" THEN
       "LPMLV30_ConfigureDisabledStates"(HoldingDisable := TRUE,
                               HeldDisable := TRUE,
                               UnholdingDisable := TRUE,
                               SuspendingDisable := FALSE,
                               SuspendedDisable := FALSE,
                               UnsuspendingDisable := FALSE,
                               CompletingDisable := TRUE,
                               CompleteDisable := TRUE,
                               disabledStates => "PackMLCfg".Cfg.disabledStatesInUnitModes["LPMLV30_MODE_PRODUCTION"]);
   END_IF;
   IF "FirstScan" THEN
       "LPMLV30_ConfigureDisabledStates"(HoldingDisable := TRUE,
                               HeldDisable := TRUE,
                               UnholdingDisable := TRUE,
                               SuspendingDisable := TRUE,
                               SuspendedDisable := TRUE,
                               UnsuspendingDisable := TRUE,
                               CompletingDisable := TRUE,
                               CompleteDisable := TRUE,
                               disabledStates => "PackMLCfg".Cfg.disabledStatesInUnitModes["LPMLV30_MODE_MANUAL"]);
   END_IF;
END_REGION

REGION Network 5: Call the EM00 Logic - xx Section
   RUNG wire#powerrail
      I_Contact( "PackMLCfg".disable.EM00.EM )
      wire#w1
      "InstEM00_00_Main"()
      Coil( "EM00".PackML_Sts.Unit.moduleActive )
   END_RUNG
   RUNG wire#powerrail
      Contact( "FirstScan" )
   END_RUNG wire#w1
   // the same network as SCL:
   "InstEM00_00_Main"(EN := NOT "PackMLCfg".disable.EM00.EM OR "FirstScan", ENO => #_w1);   // "EM00_00_Main"
   "EM00".PackML_Sts.Unit.moduleActive := #_w1;
END_REGION

REGION Network 6: Call the EM01 Logic - xx Section
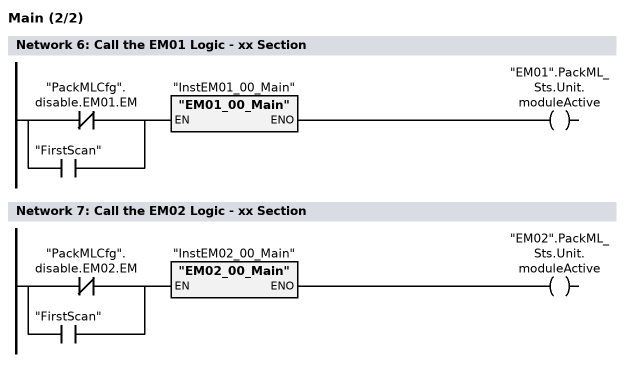
   RUNG wire#powerrail
      I_Contact( "PackMLCfg".disable.EM01.EM )
      wire#w1
      "InstEM01_00_Main"()
      Coil( "EM01".PackML_Sts.Unit.moduleActive )
   END_RUNG
   RUNG wire#powerrail
      Contact( "FirstScan" )
   END_RUNG wire#w1
   // the same network as SCL:
   "InstEM01_00_Main"(EN := NOT "PackMLCfg".disable.EM01.EM OR "FirstScan", ENO => #_w1);   // "EM01_00_Main"
   "EM01".PackML_Sts.Unit.moduleActive := #_w1;
END_REGION

REGION Network 7: Call the EM02 Logic - xx Section
   RUNG wire#powerrail
      I_Contact( "PackMLCfg".disable.EM02.EM )
      wire#w1
      "InstEM02_00_Main"()
      Coil( "EM02".PackML_Sts.Unit.moduleActive )
   END_RUNG
   RUNG wire#powerrail
      Contact( "FirstScan" )
   END_RUNG wire#w1
   // the same network as SCL:
   "InstEM02_00_Main"(EN := NOT "PackMLCfg".disable.EM02.EM OR "FirstScan", ENO => #_w1);   // "EM02_00_Main"
   "EM02".PackML_Sts.Unit.moduleActive := #_w1;
END_REGION
END_ORGANIZATION_BLOCK

// folder: EM00_Transport

FUNCTION_BLOCK "EM00_CM06_Conveyor"   // FB2, LAD
TITLE = EM00_CM04
{ S7_Optimized_Access := 'TRUE' }
AUTHOR : tech.team.motioncontrol@siemens.com
FAMILY : CPG
VERSION : 1.1
// Support: tech.team.motioncontrol@siemens.com
   VAR
      statDummyBool : Bool;   // dummy bool - placeholder
   END_VAR
BEGIN

REGION Network 1: *** Begin the Setpoint Management Information Section ***
END_REGION

REGION Network 2: *** Begin the Logic Section ***
END_REGION

REGION Network 3: *** Begin the Event Information Section ***
END_REGION

REGION Network 4: *** Begin the State Model Status Feedback Section ***
END_REGION

REGION Network 5: *** Call the PackML Module Initialize Logic ***
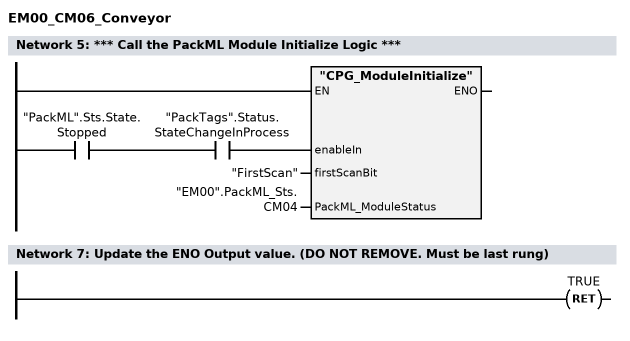
   RUNG wire#powerrail
      "CPG_ModuleInitialize"(enableIn := wire#w1, firstScanBit := "FirstScan", PackML_ModuleStatus := "EM00".PackML_Sts.CM04)
   END_RUNG
   RUNG wire#powerrail
      Contact( "PackML".Sts.State.Stopped )
      Contact( "PackTags".Status.StateChangeInProcess )
   END_RUNG wire#w1
   // the same network as SCL:
   "CPG_ModuleInitialize"(enableIn := "PackML".Sts.State.Stopped AND "PackTags".Status.StateChangeInProcess,
                          firstScanBit := "FirstScan",
                          PackML_ModuleStatus := "EM00".PackML_Sts.CM04);
END_REGION

REGION Network 7: Update the ENO Output value. (DO NOT REMOVE. Must be last rung)
   RUNG wire#powerrail
      ReturnCoil( TRUE )
   END_RUNG
   // the same network as SCL:
   ENO := TRUE;
   RETURN;
END_REGION
END_FUNCTION_BLOCK

FUNCTION_BLOCK "EM00_00_Main"   // FB31640, LAD
TITLE = EM00_00_Main
{ S7_Optimized_Access := 'TRUE' }
AUTHOR : tech.team.motioncontrol@siemens.com
FAMILY : CPG
VERSION : 1.1
// Support: tech.team.motioncontrol@siemens.com
   VAR
      instEventControl : "EM00_01_EventControl";   // Instance DB - EM's Event Control Logic
      instPackML_ModuleSum : "EM00_02_PackML_ModuleSum";   // Instance DB - EM's PackML Module Summation Logic
      instCM01 : "EM00_CM01_MainOpStation";   // Instance DB - CM01
      instCM02 : "EM00_CM02_Conveyor";   // Instance DB - CM02
      instCM03 : "EM00_CM03_ConveyorCrossing";   // Instance DB - CM03
      instCM04 : "EM00_CM04_Conveyor";   // Instance DB - CM04
      instCM05 : "EM00_CM05_ConveyorCrossing";   // Instance DB - CM05
   END_VAR
   VAR_TEMP   // added for the SCL form of the ladder/FBD networks
      _w1 : Bool;
   END_VAR
BEGIN

REGION Network 1: *** BEGIN MAIN LOGIC SECTION ***
END_REGION

REGION Network 2: Call the Control Module Logic - Main Oper. Station